(* Logix 5000 project; controller PLC_MCC1201_220AP1 vendor 1 type 14 code 164 rev 35.11; software revision 35.00; part 21 of 25 *)
(* tags used below, declared in another part *)
   GP_M225_AccessArea_FarSide : GP_AccessArea;
   GP_M225_AccessArea_FarSide_STC : GP_AccessArea_STC;
   GP_M225_AccessArea_OpSide : GP_AccessArea;
   GP_M225_AccessArea_OpSide_STC : GP_AccessArea_STC;
   TMP_xDummy : BOOL;
   xDebugOFF : BOOL;
   AFI : ALIAS FOR B3[7].15;
   GP_OB_InitializeMain : GP_OB_Initialize;
   M203DROP : MAC_DROPCONV;
   M203DROP_HMR : MAC_DROPCONV_HMR;
   M203DROP_HMW : MAC_DROPCONV_HMW;
   M205BREAKER : MAC_BREAKER;
   M205BREAKER_ALM : MAC_BREAKER_ALM;
   M205BREAKER_HMR : MAC_BREAKER_HMR;
   M205BREAKER_HMW : MAC_BREAKER_HMW;
   M225 : MAC_EMERGENCYXCUT;
   M225S_AOI_AccessArea : STRUCT_AccessArea;
   N54 : DINT[501];
   Status : INT;   // INT tag to retrieve Status value through GSV created during conversion
   TMP_xAlwaysOFF : BOOL;
   Z200 : MAC_Zone_ML;
   Z200_UPS : ZONE_UPS;
(* MainProgram, continued *)

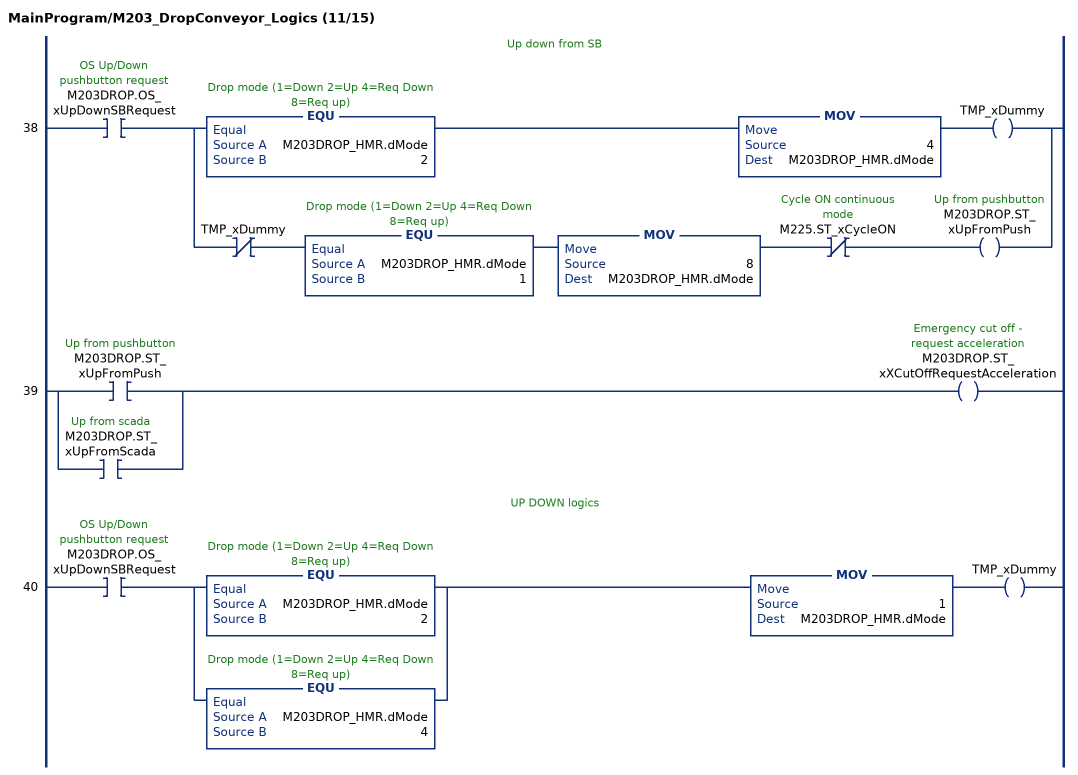
   [picture p354: MainProgram/M203_DropConveyor_Logics rungs 38-40]
   // Up down from SB
   38: XIC(M203DROP.OS_xUpDownSBRequest)[EQU(M203DROP_HMR.dMode,2) MOV(4,M203DROP_HMR.dMode) OTE(TMP_xDummy) ,XIO(TMP_xDummy) EQU(M203DROP_HMR.dMode,1) MOV(8,M203DROP_HMR.dMode) XIO(M225.ST_xCycleON) OTE(M203DROP.ST_xUpFromPush) ];
   39: [XIC(M203DROP.ST_xUpFromPush) ,XIC(M203DROP.ST_xUpFromScada) ]OTE(M203DROP.ST_xXCutOffRequestAcceleration);
   // UP DOWN logics
   40: XIC(M203DROP.OS_xUpDownSBRequest)[EQU(M203DROP_HMR.dMode,2) ,EQU(M203DROP_HMR.dMode,4) ]MOV(1,M203DROP_HMR.dMode)OTE(TMP_xDummy);
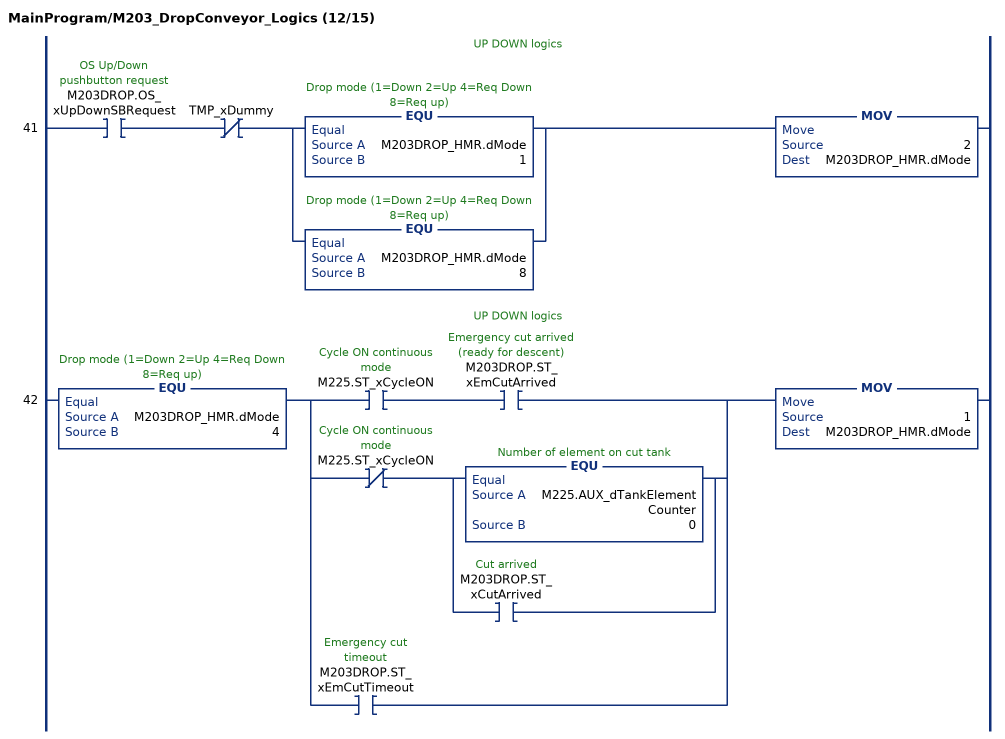
   // UP DOWN logics
   41: XIC(M203DROP.OS_xUpDownSBRequest)XIO(TMP_xDummy)[EQU(M203DROP_HMR.dMode,1) ,EQU(M203DROP_HMR.dMode,8) ]MOV(2,M203DROP_HMR.dMode);
   // UP DOWN logics
   42: EQU(M203DROP_HMR.dMode,4)[XIC(M225.ST_xCycleON) XIC(M203DROP.ST_xEmCutArrived) ,XIO(M225.ST_xCycleON) [EQU(M225.AUX_dTankElementCounter,0) ,XIC(M203DROP.ST_xCutArrived) ] ,XIC(M203DROP.ST_xEmCutTimeout) ]MOV(1,M203DROP_HMR.dMode);
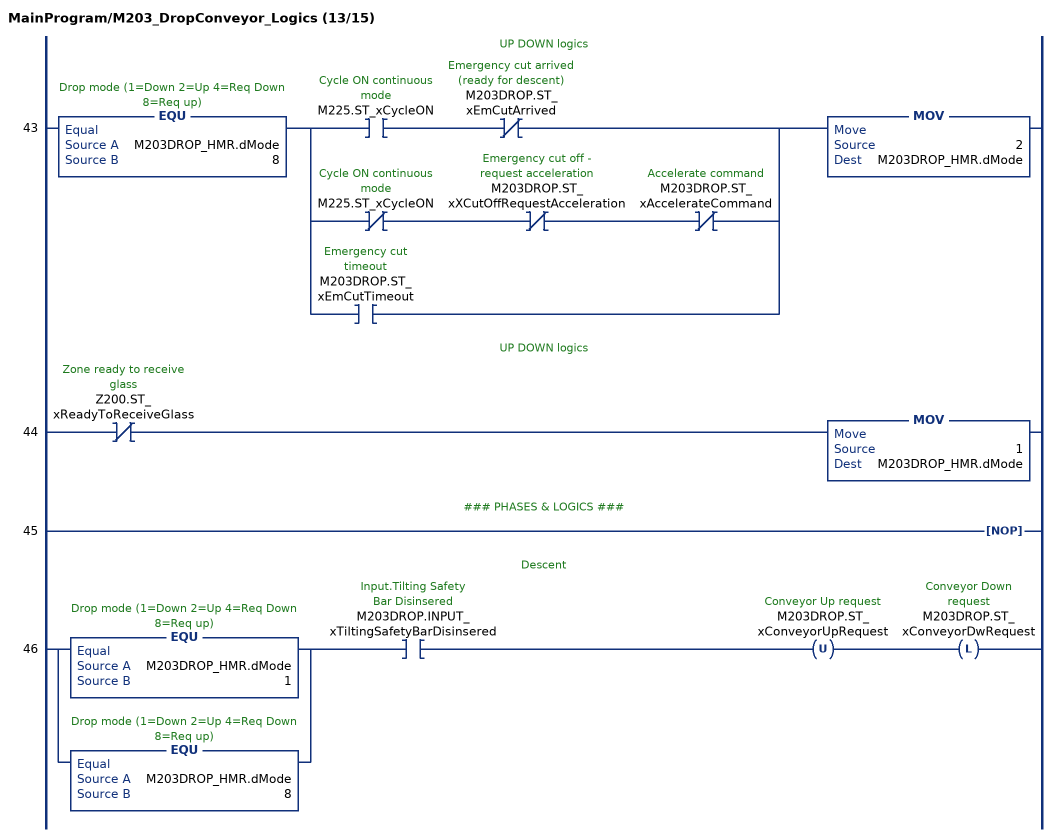
   // UP DOWN logics
   43: EQU(M203DROP_HMR.dMode,8)[XIC(M225.ST_xCycleON) XIO(M203DROP.ST_xEmCutArrived) ,XIO(M225.ST_xCycleON) XIO(M203DROP.ST_xXCutOffRequestAcceleration) XIO(M203DROP.ST_xAccelerateCommand) ,XIC(M203DROP.ST_xEmCutTimeout) ]MOV(2,M203DROP_HMR.dMode);
   // UP DOWN logics
   44: XIO(Z200.ST_xReadyToReceiveGlass)MOV(1,M203DROP_HMR.dMode);
   // ### PHASES & LOGICS ###
   45: NOP();
   // Descent
   46: [EQU(M203DROP_HMR.dMode,1) ,EQU(M203DROP_HMR.dMode,8) ]XIC(M203DROP.INPUT_xTiltingSafetyBarDisinsered)OTU(M203DROP.ST_xConveyorUpRequest)OTL(M203DROP.ST_xConveyorDwRequest);
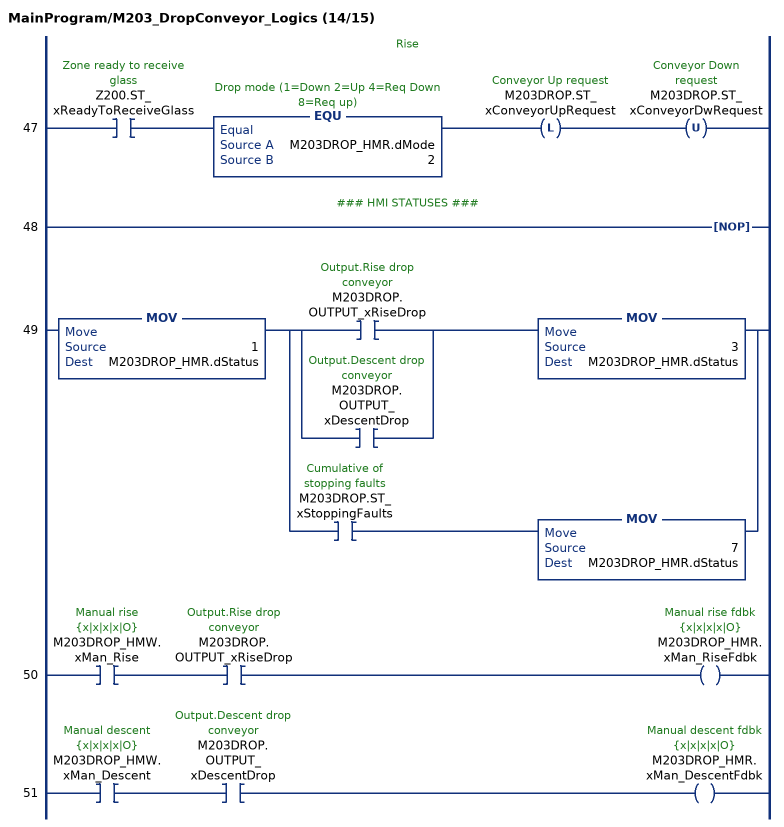
   // Rise
   47: XIC(Z200.ST_xReadyToReceiveGlass)EQU(M203DROP_HMR.dMode,2)OTL(M203DROP.ST_xConveyorUpRequest)OTU(M203DROP.ST_xConveyorDwRequest);
   // ### HMI STATUSES ###
   48: NOP();
   49: MOV(1,M203DROP_HMR.dStatus)[[XIC(M203DROP.OUTPUT_xRiseDrop) ,XIC(M203DROP.OUTPUT_xDescentDrop) ] MOV(3,M203DROP_HMR.dStatus) ,XIC(M203DROP.ST_xStoppingFaults) MOV(7,M203DROP_HMR.dStatus) ];
   50: XIC(M203DROP_HMW.xMan_Rise)XIC(M203DROP.OUTPUT_xRiseDrop)OTE(M203DROP_HMR.xMan_RiseFdbk);
   51: XIC(M203DROP_HMW.xMan_Descent)XIC(M203DROP.OUTPUT_xDescentDrop)OTE(M203DROP_HMR.xMan_DescentFdbk);
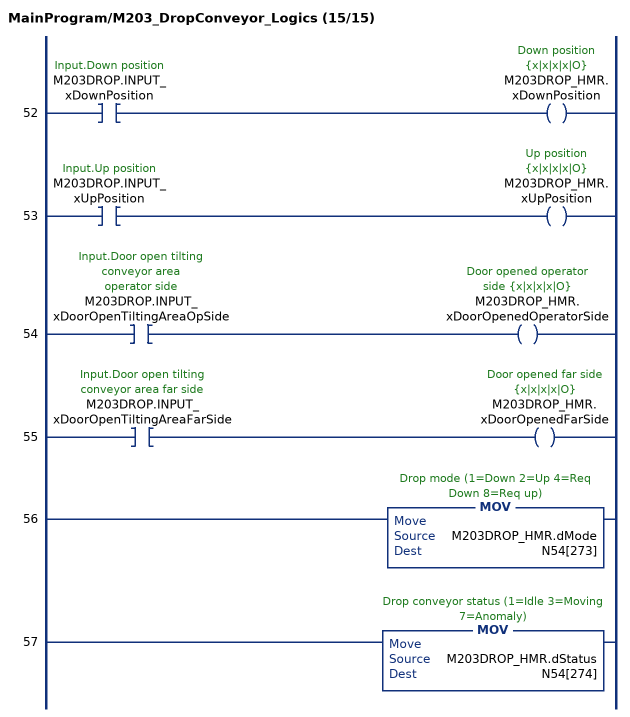
   52: XIC(M203DROP.INPUT_xDownPosition)OTE(M203DROP_HMR.xDownPosition);
   53: XIC(M203DROP.INPUT_xUpPosition)OTE(M203DROP_HMR.xUpPosition);
   54: XIC(M203DROP.INPUT_xDoorOpenTiltingAreaOpSide)OTE(M203DROP_HMR.xDoorOpenedOperatorSide);
   55: XIC(M203DROP.INPUT_xDoorOpenTiltingAreaFarSide)OTE(M203DROP_HMR.xDoorOpenedFarSide);
   56: MOV(M203DROP_HMR.dMode,N54[273]);
   57: MOV(M203DROP_HMR.dStatus,N54[274]);
END_ROUTINE

ROUTINE M205B_Breaker_Faults   (* ladder *)
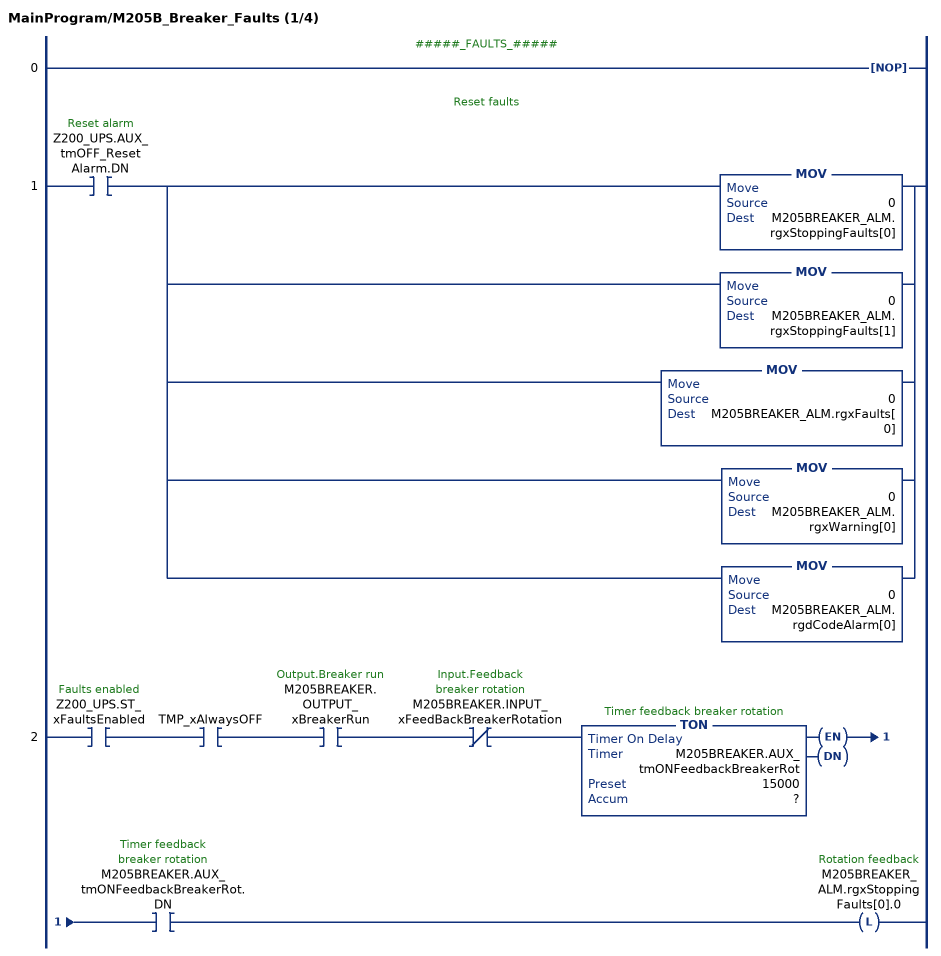
   // #####_FAULTS_#####
   0: NOP();
   // Reset faults
   1: XIC(Z200_UPS.AUX_tmOFF_ResetAlarm.DN)[MOV(0,M205BREAKER_ALM.rgxStoppingFaults[0]) ,MOV(0,M205BREAKER_ALM.rgxStoppingFaults[1]) ,MOV(0,M205BREAKER_ALM.rgxFaults[0]) ,MOV(0,M205BREAKER_ALM.rgxWarning[0]) ,MOV(0,M205BREAKER_ALM.rgdCodeAlarm[0]) ];
   2: XIC(Z200_UPS.ST_xFaultsEnabled)XIC(TMP_xAlwaysOFF)XIC(M205BREAKER.OUTPUT_xBreakerRun)XIO(M205BREAKER.INPUT_xFeedBackBreakerRotation)TON(M205BREAKER.AUX_tmONFeedbackBreakerRot,?,?)XIC(M205BREAKER.AUX_tmONFeedbackBreakerRot.DN)OTL(M205BREAKER_ALM.rgxStoppingFaults[0].0);
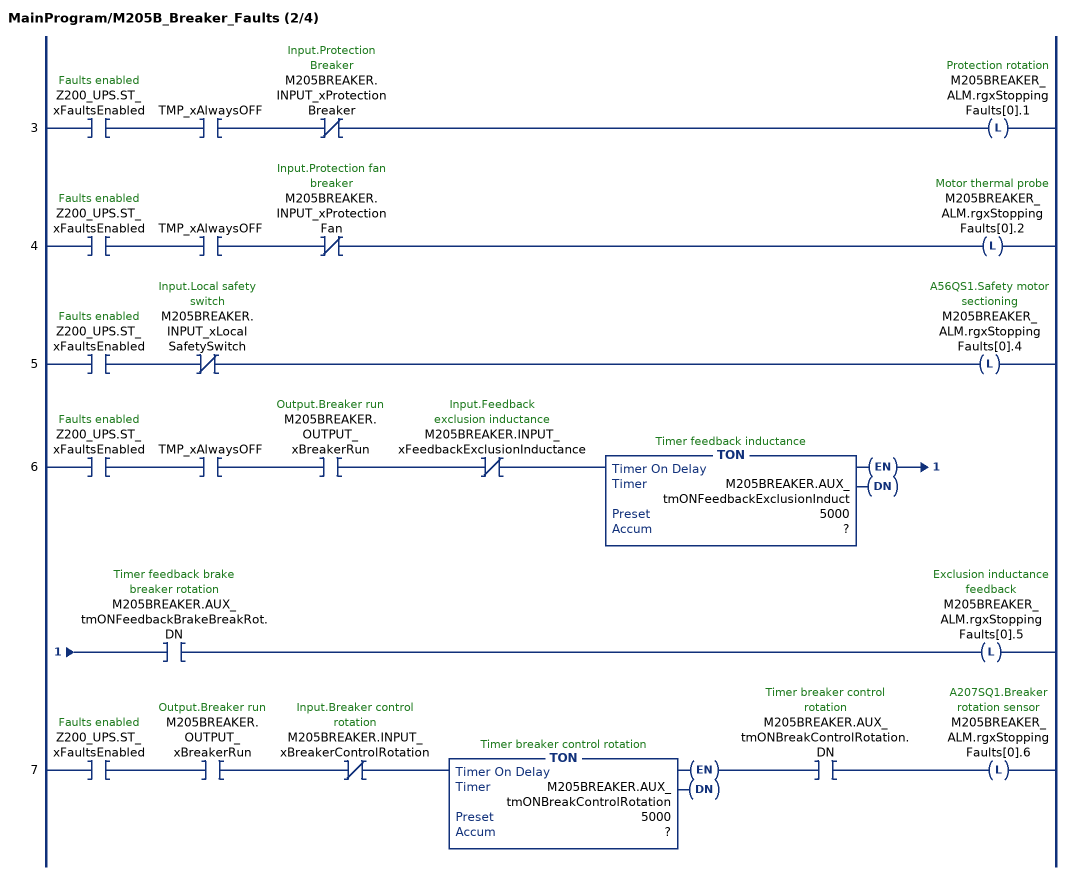
   3: XIC(Z200_UPS.ST_xFaultsEnabled)XIC(TMP_xAlwaysOFF)XIO(M205BREAKER.INPUT_xProtectionBreaker)OTL(M205BREAKER_ALM.rgxStoppingFaults[0].1);
   4: XIC(Z200_UPS.ST_xFaultsEnabled)XIC(TMP_xAlwaysOFF)XIO(M205BREAKER.INPUT_xProtectionFan)OTL(M205BREAKER_ALM.rgxStoppingFaults[0].2);
   5: XIC(Z200_UPS.ST_xFaultsEnabled)XIO(M205BREAKER.INPUT_xLocalSafetySwitch)OTL(M205BREAKER_ALM.rgxStoppingFaults[0].4);
   6: XIC(Z200_UPS.ST_xFaultsEnabled)XIC(TMP_xAlwaysOFF)XIC(M205BREAKER.OUTPUT_xBreakerRun)XIO(M205BREAKER.INPUT_xFeedbackExclusionInductance)TON(M205BREAKER.AUX_tmONFeedbackExclusionInduct,?,?)XIC(M205BREAKER.AUX_tmONFeedbackBrakeBreakRot.DN)OTL(M205BREAKER_ALM.rgxStoppingFaults[0].5);
   7: XIC(Z200_UPS.ST_xFaultsEnabled)XIC(M205BREAKER.OUTPUT_xBreakerRun)XIO(M205BREAKER.INPUT_xBreakerControlRotation)TON(M205BREAKER.AUX_tmONBreakControlRotation,?,?)XIC(M205BREAKER.AUX_tmONBreakControlRotation.DN)OTL(M205BREAKER_ALM.rgxStoppingFaults[0].6);
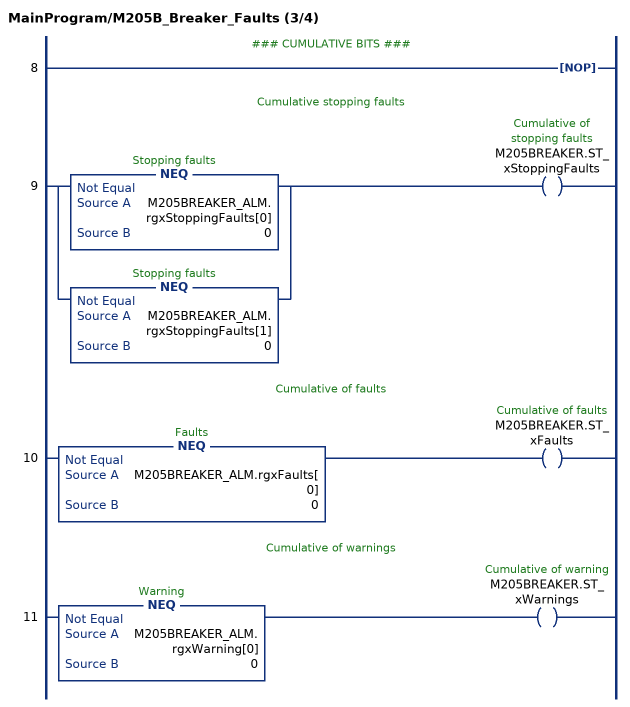
   // ### CUMULATIVE BITS ###
   8: NOP();
   // Cumulative stopping faults
   9: [NEQ(M205BREAKER_ALM.rgxStoppingFaults[0],0) ,NEQ(M205BREAKER_ALM.rgxStoppingFaults[1],0) ]OTE(M205BREAKER.ST_xStoppingFaults);
   // Cumulative of faults
   10: NEQ(M205BREAKER_ALM.rgxFaults[0],0)OTE(M205BREAKER.ST_xFaults);
   // Cumulative of warnings
   11: NEQ(M205BREAKER_ALM.rgxWarning[0],0)OTE(M205BREAKER.ST_xWarnings);
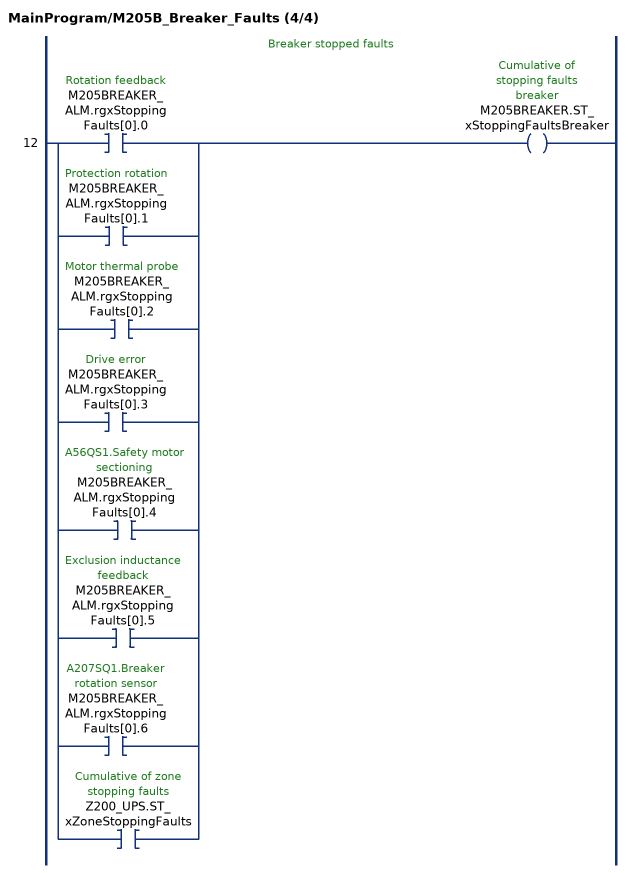
   // Breaker stopped faults
   12: [XIC(M205BREAKER_ALM.rgxStoppingFaults[0].0) ,XIC(M205BREAKER_ALM.rgxStoppingFaults[0].1) ,XIC(M205BREAKER_ALM.rgxStoppingFaults[0].2) ,XIC(M205BREAKER_ALM.rgxStoppingFaults[0].3) ,XIC(M205BREAKER_ALM.rgxStoppingFaults[0].4) ,XIC(M205BREAKER_ALM.rgxStoppingFaults[0].5) ,XIC(M205BREAKER_ALM.rgxStoppingFaults[0].6) ,XIC(Z200_UPS.ST_xZoneStoppingFaults) ]OTE(M205BREAKER.ST_xStoppingFaultsBreaker);
END_ROUTINE

ROUTINE M205B_Breaker_Logics   (* ladder *)
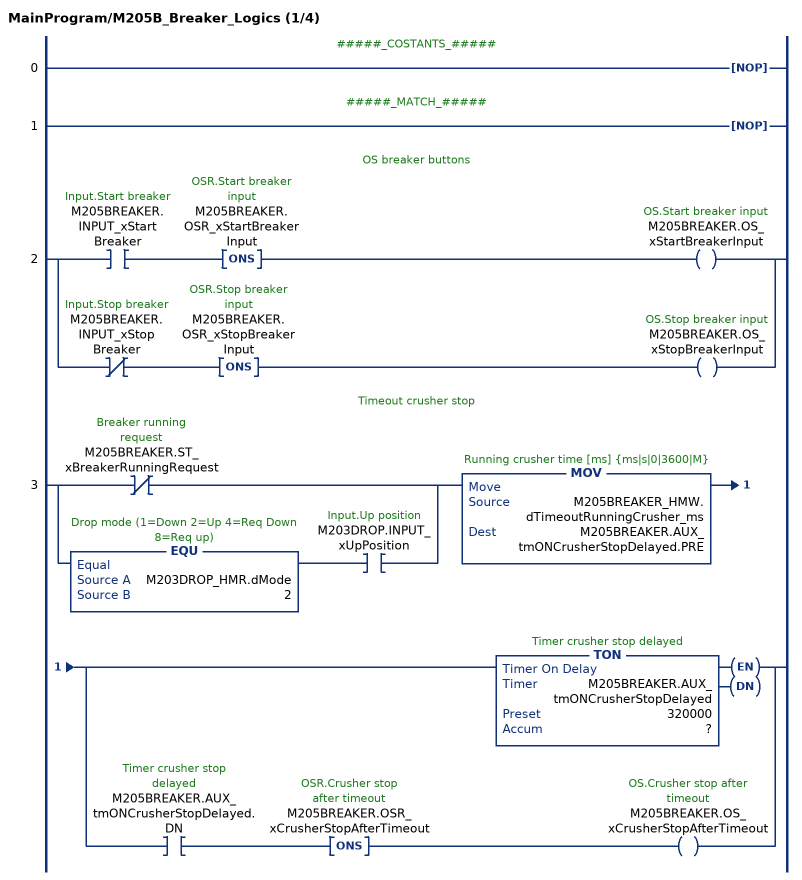
   // #####_COSTANTS_#####
   0: NOP();
   // #####_MATCH_#####
   1: NOP();
   // OS breaker buttons
   2: [XIC(M205BREAKER.INPUT_xStartBreaker) ONS(M205BREAKER.OSR_xStartBreakerInput) OTE(M205BREAKER.OS_xStartBreakerInput) ,XIO(M205BREAKER.INPUT_xStopBreaker) ONS(M205BREAKER.OSR_xStopBreakerInput) OTE(M205BREAKER.OS_xStopBreakerInput) ];
   // Timeout crusher stop
   3: [XIO(M205BREAKER.ST_xBreakerRunningRequest) ,EQU(M203DROP_HMR.dMode,2) XIC(M203DROP.INPUT_xUpPosition) ]MOV(M205BREAKER_HMW.dTimeoutRunningCrusher_ms,M205BREAKER.AUX_tmONCrusherStopDelayed.PRE)[TON(M205BREAKER.AUX_tmONCrusherStopDelayed,?,?) ,XIC(M205BREAKER.AUX_tmONCrusherStopDelayed.DN) ONS(M205BREAKER.OSR_xCrusherStopAfterTimeout) OTE(M205BREAKER.OS_xCrusherStopAfterTimeout) ];
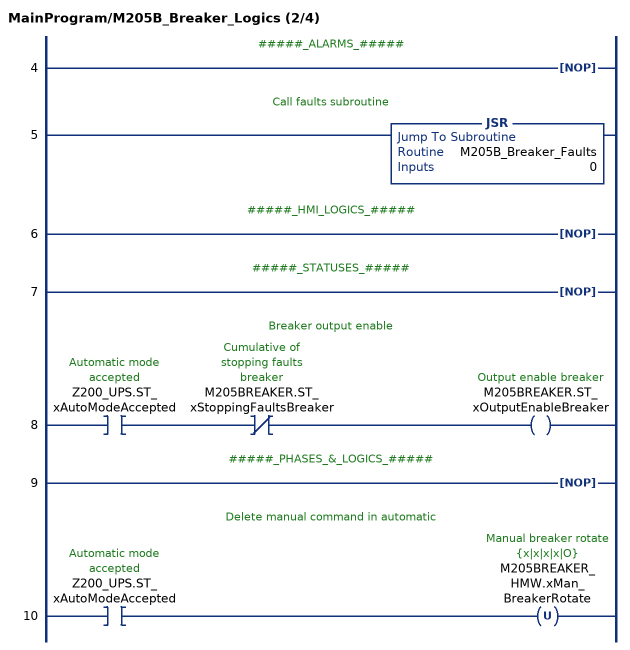
   // #####_ALARMS_#####
   4: NOP();
   // Call faults subroutine
   5: JSR(M205B_Breaker_Faults,0);
   // #####_HMI_LOGICS_#####
   6: NOP();
   // #####_STATUSES_#####
   7: NOP();
   // Breaker output enable
   8: XIC(Z200_UPS.ST_xAutoModeAccepted)XIO(M205BREAKER.ST_xStoppingFaultsBreaker)OTE(M205BREAKER.ST_xOutputEnableBreaker);
   // #####_PHASES_&_LOGICS_#####
   9: NOP();
   // Delete manual command in automatic
   10: XIC(Z200_UPS.ST_xAutoModeAccepted)OTU(M205BREAKER_HMW.xMan_BreakerRotate);
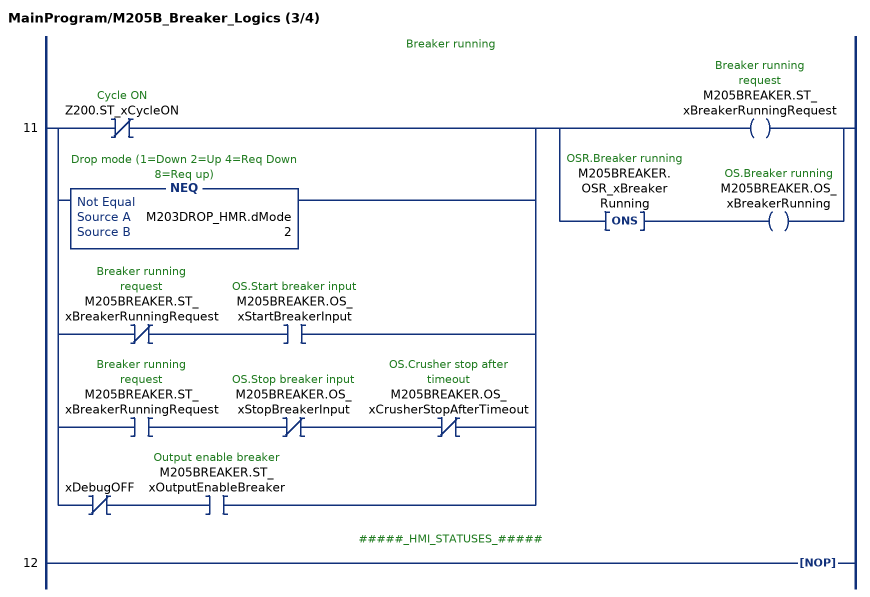
   // Breaker running
   11: [XIO(Z200.ST_xCycleON) ,NEQ(M203DROP_HMR.dMode,2) ,XIO(M205BREAKER.ST_xBreakerRunningRequest) XIC(M205BREAKER.OS_xStartBreakerInput) ,XIC(M205BREAKER.ST_xBreakerRunningRequest) XIO(M205BREAKER.OS_xStopBreakerInput) XIO(M205BREAKER.OS_xCrusherStopAfterTimeout) ,XIO(xDebugOFF) XIC(M205BREAKER.ST_xOutputEnableBreaker) ][OTE(M205BREAKER.ST_xBreakerRunningRequest) ,ONS(M205BREAKER.OSR_xBreakerRunning) OTE(M205BREAKER.OS_xBreakerRunning) ];
   // #####_HMI_STATUSES_#####
   12: NOP();
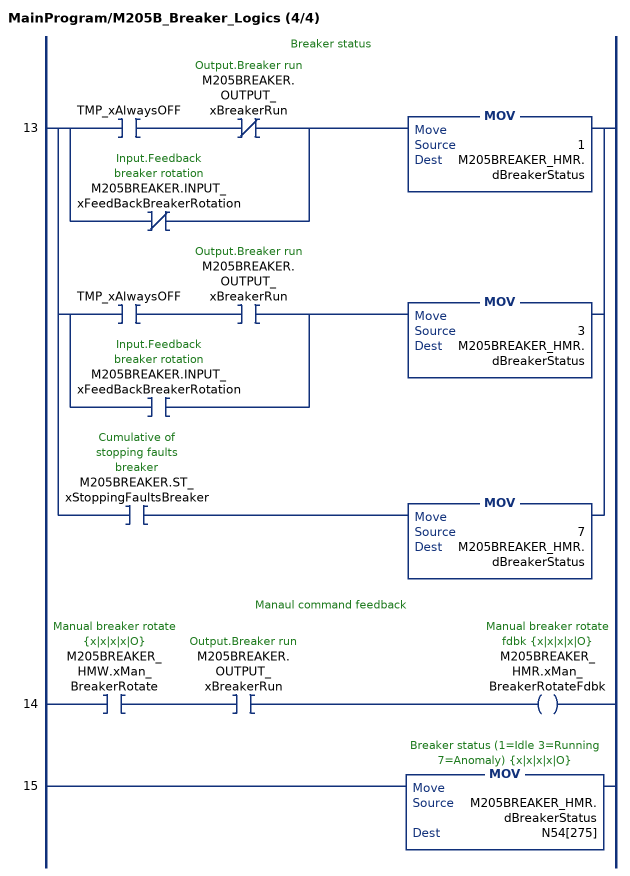
   // Breaker status
   13: [[XIC(TMP_xAlwaysOFF) XIO(M205BREAKER.OUTPUT_xBreakerRun) ,XIO(M205BREAKER.INPUT_xFeedBackBreakerRotation) ] MOV(1,M205BREAKER_HMR.dBreakerStatus) ,[XIC(TMP_xAlwaysOFF) XIC(M205BREAKER.OUTPUT_xBreakerRun) ,XIC(M205BREAKER.INPUT_xFeedBackBreakerRotation) ] MOV(3,M205BREAKER_HMR.dBreakerStatus) ,XIC(M205BREAKER.ST_xStoppingFaultsBreaker) MOV(7,M205BREAKER_HMR.dBreakerStatus) ];
   // Manaul command feedback
   14: XIC(M205BREAKER_HMW.xMan_BreakerRotate)XIC(M205BREAKER.OUTPUT_xBreakerRun)OTE(M205BREAKER_HMR.xMan_BreakerRotateFdbk);
   15: MOV(M205BREAKER_HMR.dBreakerStatus,N54[275]);
END_ROUTINE

ROUTINE M225_EmCut_AccessArea   (* ladder *)
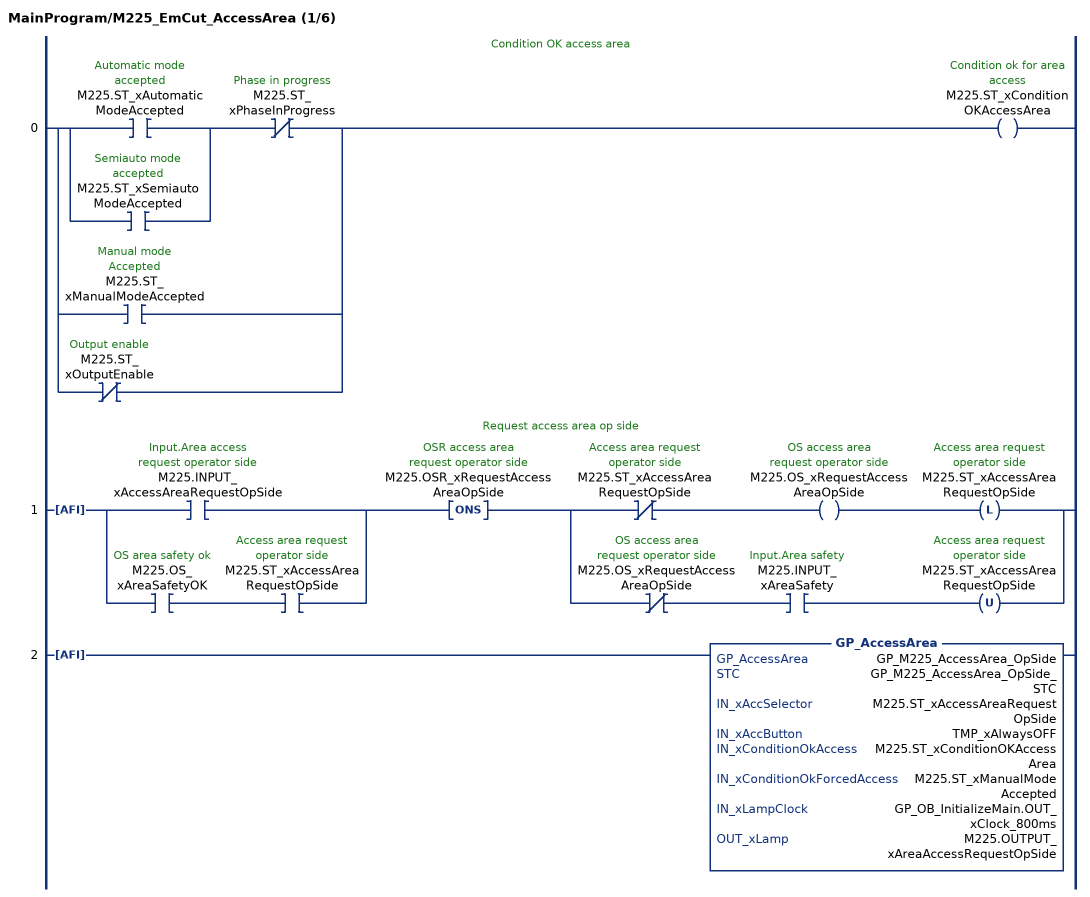
   // Condition OK access area
   0: [[XIC(M225.ST_xAutomaticModeAccepted) ,XIC(M225.ST_xSemiautoModeAccepted) ] XIO(M225.ST_xPhaseInProgress) ,XIC(M225.ST_xManualModeAccepted) ,XIO(M225.ST_xOutputEnable) ]OTE(M225.ST_xConditionOKAccessArea);
   // Request access area op side
   1: AFI()[XIC(M225.INPUT_xAccessAreaRequestOpSide) ,XIC(M225.OS_xAreaSafetyOK) XIC(M225.ST_xAccessAreaRequestOpSide) ]ONS(M225.OSR_xRequestAccessAreaOpSide)[XIO(M225.ST_xAccessAreaRequestOpSide) OTE(M225.OS_xRequestAccessAreaOpSide) OTL(M225.ST_xAccessAreaRequestOpSide) ,XIO(M225.OS_xRequestAccessAreaOpSide) XIC(M225.INPUT_xAreaSafety) OTU(M225.ST_xAccessAreaRequestOpSide) ];
   2: AFI()GP_AccessArea(GP_M225_AccessArea_OpSide,GP_M225_AccessArea_OpSide_STC,M225.ST_xAccessAreaRequestOpSide,TMP_xAlwaysOFF,M225.ST_xConditionOKAccessArea,M225.ST_xManualModeAccepted,GP_OB_InitializeMain.OUT_xClock_800ms,M225.OUTPUT_xAreaAccessRequestOpSide);
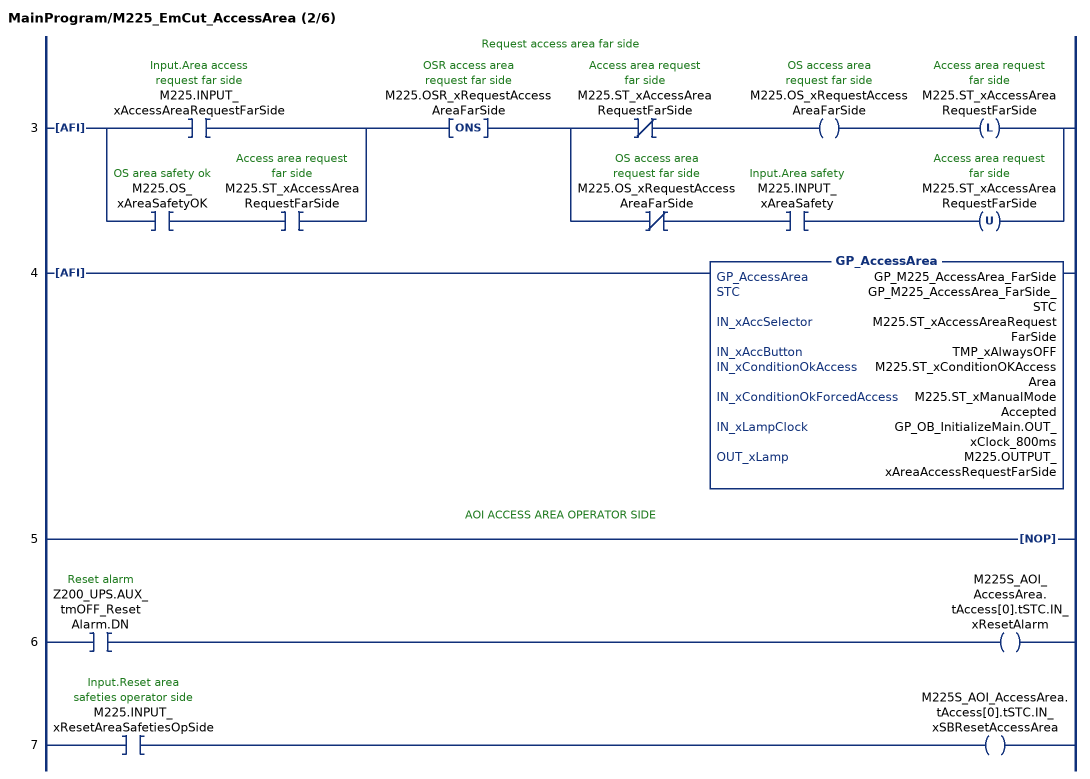
   // Request access area far side
   3: AFI()[XIC(M225.INPUT_xAccessAreaRequestFarSide) ,XIC(M225.OS_xAreaSafetyOK) XIC(M225.ST_xAccessAreaRequestFarSide) ]ONS(M225.OSR_xRequestAccessAreaFarSide)[XIO(M225.ST_xAccessAreaRequestFarSide) OTE(M225.OS_xRequestAccessAreaFarSide) OTL(M225.ST_xAccessAreaRequestFarSide) ,XIO(M225.OS_xRequestAccessAreaFarSide) XIC(M225.INPUT_xAreaSafety) OTU(M225.ST_xAccessAreaRequestFarSide) ];
   4: AFI()GP_AccessArea(GP_M225_AccessArea_FarSide,GP_M225_AccessArea_FarSide_STC,M225.ST_xAccessAreaRequestFarSide,TMP_xAlwaysOFF,M225.ST_xConditionOKAccessArea,M225.ST_xManualModeAccepted,GP_OB_InitializeMain.OUT_xClock_800ms,M225.OUTPUT_xAreaAccessRequestFarSide);
   // AOI ACCESS AREA OPERATOR SIDE
   5: NOP();
   6: XIC(Z200_UPS.AUX_tmOFF_ResetAlarm.DN)OTE(M225S_AOI_AccessArea.tAccess[0].tSTC.IN_xResetAlarm);
   7: XIC(M225.INPUT_xResetAreaSafetiesOpSide)OTE(M225S_AOI_AccessArea.tAccess[0].tSTC.IN_xSBResetAccessArea);
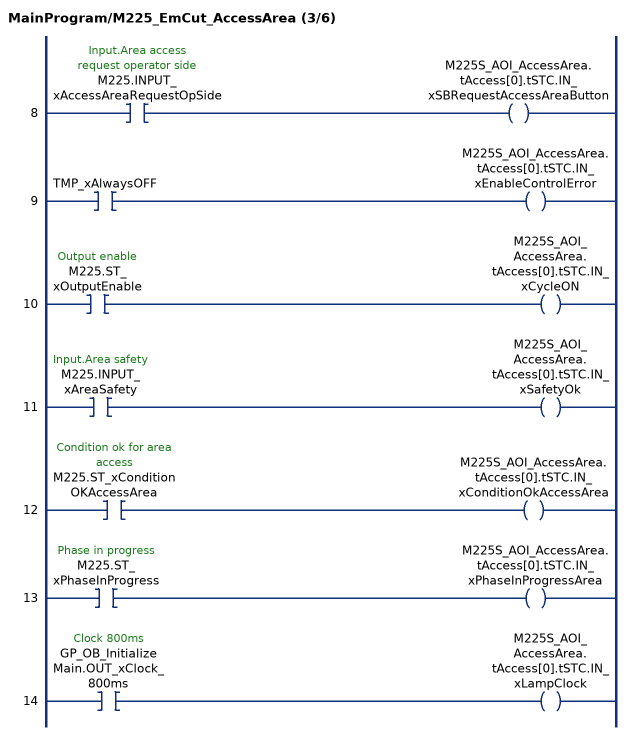
   8: XIC(M225.INPUT_xAccessAreaRequestOpSide)OTE(M225S_AOI_AccessArea.tAccess[0].tSTC.IN_xSBRequestAccessAreaButton);
   9: XIC(TMP_xAlwaysOFF)OTE(M225S_AOI_AccessArea.tAccess[0].tSTC.IN_xEnableControlError);
   10: XIC(M225.ST_xOutputEnable)OTE(M225S_AOI_AccessArea.tAccess[0].tSTC.IN_xCycleON);
   11: XIC(M225.INPUT_xAreaSafety)OTE(M225S_AOI_AccessArea.tAccess[0].tSTC.IN_xSafetyOk);
   12: XIC(M225.ST_xConditionOKAccessArea)OTE(M225S_AOI_AccessArea.tAccess[0].tSTC.IN_xConditionOkAccessArea);
   13: XIC(M225.ST_xPhaseInProgress)OTE(M225S_AOI_AccessArea.tAccess[0].tSTC.IN_xPhaseInProgressArea);
   14: XIC(GP_OB_InitializeMain.OUT_xClock_800ms)OTE(M225S_AOI_AccessArea.tAccess[0].tSTC.IN_xLampClock);
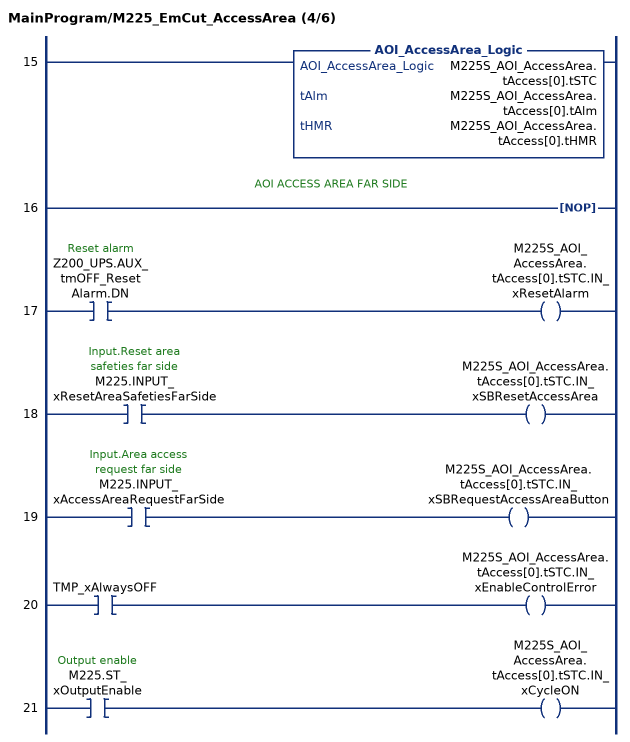
   15: AOI_AccessArea_Logic(M225S_AOI_AccessArea.tAccess[0].tSTC,M225S_AOI_AccessArea.tAccess[0].tAlm,M225S_AOI_AccessArea.tAccess[0].tHMR);
   // AOI ACCESS AREA FAR SIDE
   16: NOP();
   17: XIC(Z200_UPS.AUX_tmOFF_ResetAlarm.DN)OTE(M225S_AOI_AccessArea.tAccess[0].tSTC.IN_xResetAlarm);
   18: XIC(M225.INPUT_xResetAreaSafetiesFarSide)OTE(M225S_AOI_AccessArea.tAccess[0].tSTC.IN_xSBResetAccessArea);
   19: XIC(M225.INPUT_xAccessAreaRequestFarSide)OTE(M225S_AOI_AccessArea.tAccess[0].tSTC.IN_xSBRequestAccessAreaButton);
   20: XIC(TMP_xAlwaysOFF)OTE(M225S_AOI_AccessArea.tAccess[0].tSTC.IN_xEnableControlError);
   21: XIC(M225.ST_xOutputEnable)OTE(M225S_AOI_AccessArea.tAccess[0].tSTC.IN_xCycleON);
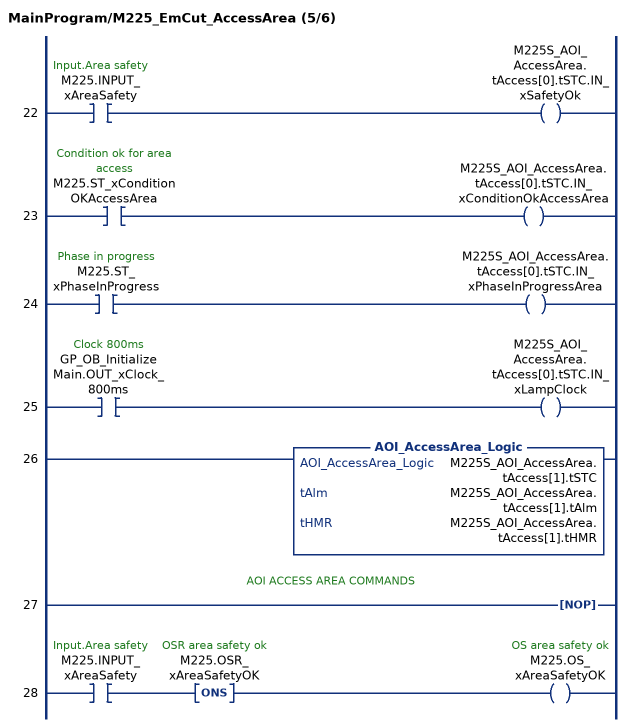
   22: XIC(M225.INPUT_xAreaSafety)OTE(M225S_AOI_AccessArea.tAccess[0].tSTC.IN_xSafetyOk);
   23: XIC(M225.ST_xConditionOKAccessArea)OTE(M225S_AOI_AccessArea.tAccess[0].tSTC.IN_xConditionOkAccessArea);
   24: XIC(M225.ST_xPhaseInProgress)OTE(M225S_AOI_AccessArea.tAccess[0].tSTC.IN_xPhaseInProgressArea);
   25: XIC(GP_OB_InitializeMain.OUT_xClock_800ms)OTE(M225S_AOI_AccessArea.tAccess[0].tSTC.IN_xLampClock);
   26: AOI_AccessArea_Logic(M225S_AOI_AccessArea.tAccess[1].tSTC,M225S_AOI_AccessArea.tAccess[1].tAlm,M225S_AOI_AccessArea.tAccess[1].tHMR);
   // AOI ACCESS AREA COMMANDS
   27: NOP();
   28: XIC(M225.INPUT_xAreaSafety)ONS(M225.OSR_xAreaSafetyOK)OTE(M225.OS_xAreaSafetyOK);
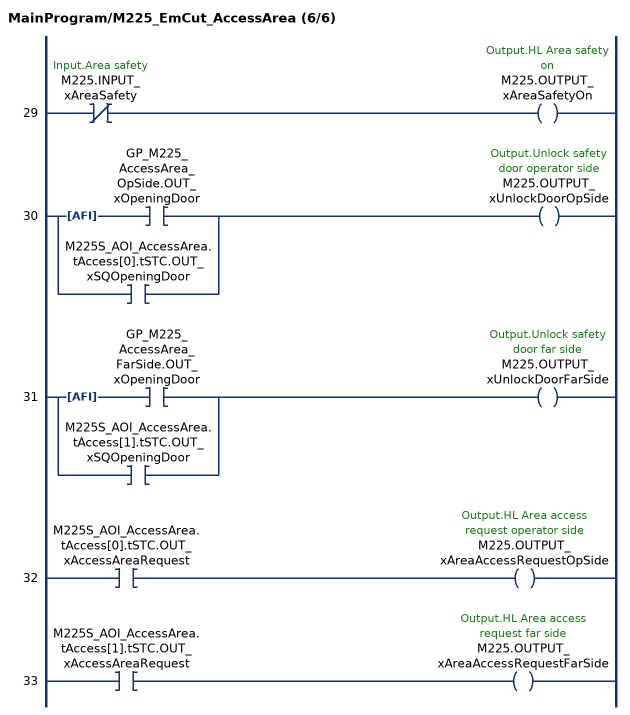
   29: XIO(M225.INPUT_xAreaSafety)OTE(M225.OUTPUT_xAreaSafetyOn);
   30: [AFI() XIC(GP_M225_AccessArea_OpSide.OUT_xOpeningDoor) ,XIC(M225S_AOI_AccessArea.tAccess[0].tSTC.OUT_xSQOpeningDoor) ]OTE(M225.OUTPUT_xUnlockDoorOpSide);
   31: [AFI() XIC(GP_M225_AccessArea_FarSide.OUT_xOpeningDoor) ,XIC(M225S_AOI_AccessArea.tAccess[1].tSTC.OUT_xSQOpeningDoor) ]OTE(M225.OUTPUT_xUnlockDoorFarSide);
   32: XIC(M225S_AOI_AccessArea.tAccess[0].tSTC.OUT_xAccessAreaRequest)OTE(M225.OUTPUT_xAreaAccessRequestOpSide);
   33: XIC(M225S_AOI_AccessArea.tAccess[1].tSTC.OUT_xAccessAreaRequest)OTE(M225.OUTPUT_xAreaAccessRequestFarSide);
END_ROUTINE
